DATA_BLOCK "2062_Warning_Data"   // DB2062
{ S7_Optimized_Access := 'FALSE' }
VERSION : 0.1
   VAR
      BTCS_WARNING_WORD_01 : Word;
      BTCS_WARNING_WORD_02 : Word;
      BTCS_WARNING_WORD_03 : Word;
      BTCS_WARNING_WORD_04 : Word;
      BTCS_WARNING_WORD_05 : Word;
      BTCS_WARNING_WORD_06 : Word;
      BTCS_WARNING_WORD_07 : Word;
      BTCS_WARNING_WORD_08 : Word;
      BTCS_WARNING_WORD_09 : Word;
      BTCS_WARNING_WORD_10 : Word;
      BTCS_WARNING_WORD_11 : Word;
      WARNING_PRSNT : Bool;
      "Alarm Tank FPT" : Bool;
      "Alarm Tank P1" : Bool;
      "Alarm Tank S1" : Bool;
      "Alarm Tank P2" : Bool;
      "Alarm Tank S2" : Bool;
      "Alarm Tank P3" : Bool;
      "Alarm Tank S3" : Bool;
      "Alarm Tank P4" : Bool;
      "Alarm Tank S4" : Bool;
      "Alarm Tank P5" : Bool;
      "Alarm Tank S5" : Bool;
      "Alarm Tank P6" : Bool;
      "Alarm Tank S6" : Bool;
      "Alarm Tank APT" : Bool;
      "LS425 FPT Level HIHI" : TON_TIME;
      "LS425 1 Port Level HIHI" : TON_TIME;
      "LS425 1 Starboard Level HIHI" : TON_TIME;
      "PS436 RIO1 Tank Group Pressure HIHI" : TON_TIME;
      "LS425 2 Port Level HIHI" : TON_TIME;
      "LS425 2 Starboard Level HIHI" : TON_TIME;
      "PS436 RIO2 Tank Group Pressure HIHI" : TON_TIME;
      "LS425 3 Port Level HIHI" : TON_TIME;
      "LS425 3 Starboard Level HIHI" : TON_TIME;
      "PS436 RIO3 Tank Group Pressure HIHI" : TON_TIME;
      "LS425 4 Port Level HIHI" : TON_TIME;
      "LS425 4 Starboard Level HIHI" : TON_TIME;
      "PS436 RIO4 Tank Group Pressure HIHI" : TON_TIME;
      "LS425 5 Port Level HIHI" : TON_TIME;
      "LS425 5 Starboard Level HIHI" : TON_TIME;
      "PS436 RIO5 Tank Group Pressure HIHI" : TON_TIME;
      "LS425 6 Port Level HIHI" : TON_TIME;
      "LS425 6 Starboard Level HIHI" : TON_TIME;
      "PS436 RIO6 Tank Group Pressure HIHI" : TON_TIME;
      "LS425 APT Level HIHI" : TON_TIME;
      "PS436 RIO7 Tank Group Pressure HIHI" : TON_TIME;
      "Water Level Override FPT" : Bool;
      "Water Level Override 1P" : Bool;
      "Water Level Override 1S" : Bool;
      "Water Level Override 2P" : Bool;
      "Water Level Override 2S" : Bool;
      "Water Level Override 3P" : Bool;
      "Water Level Override 3S" : Bool;
      "Water Level Override 4P" : Bool;
      "Water Level Override 4S" : Bool;
      "Water Level Override 5P" : Bool;
      "Water Level Override 5S" : Bool;
      "Water Level Override 6P" : Bool;
      "Water Level Override 6S" : Bool;
      "Water Level Override APT" : Bool;
      BTCS_WARNING_WORD_12 : Word;
      BTCS_WARNING_WORD_13 : Word;
      BTCS_WARNING_WORD_14 : Word;
      BTCS_WARNING_WORD_15 : Word;
      BTCS_WARNING_WORD_16 : Word;
      BTCS_WARNING_WORD_17 : Word;
      BTCS_WARNING_WORD_18 : Word;
      "Water Level Override" : Bool;
      "Water Level Override_flag" : Bool;
      "Water Level Override_Aux" : Bool;
   END_VAR
BEGIN
   "LS425 2 Port Level HIHI".PT := T#10s;
   "LS425 2 Starboard Level HIHI".PT := T#10s;
   "PS436 RIO2 Tank Group Pressure HIHI".PT := T#3s;
   "LS425 FPT Level HIHI".PT := T#10s;
   "LS425 1 Port Level HIHI".PT := T#10s;
   "LS425 1 Starboard Level HIHI".PT := T#3s;
END_DATA_BLOCK

DATA_BLOCK "503_WARNING CHCK_DB_2063"   // DB2063
{ S7_Optimized_Access := 'TRUE' }
VERSION : 0.1
// stored: InstanceOfName 503_ALARM CHCK
"503_ALARM CHCK"
BEGIN
END_DATA_BLOCK

DATA_BLOCK "FIT418_2P_ALM_ANALOG_DB"   // DB2064
{ S7_Optimized_Access := 'FALSE' }
VERSION : 0.1
// stored: InstanceOfName 502_ALM_ANALOG
"502_ALM_ANALOG"
BEGIN
END_DATA_BLOCK

DATA_BLOCK "FIT420PORT_ALM_ANALOG_DB"   // DB2065
{ S7_Optimized_Access := 'FALSE' }
VERSION : 0.1
// stored: InstanceOfName 502_ALM_ANALOG
"502_ALM_ANALOG"
BEGIN
END_DATA_BLOCK

DATA_BLOCK "FIT417_2S_ALM_ANALOG_DB"   // DB2066
{ S7_Optimized_Access := 'FALSE' }
VERSION : 0.1
// stored: InstanceOfName 502_ALM_ANALOG
"502_ALM_ANALOG"
BEGIN
END_DATA_BLOCK

DATA_BLOCK "FIT419_ALM_ANALOG_DB"   // DB2067
{ S7_Optimized_Access := 'FALSE' }
VERSION : 0.1
// stored: InstanceOfName 502_ALM_ANALOG
"502_ALM_ANALOG"
BEGIN
END_DATA_BLOCK

DATA_BLOCK "2068_Sys_Status_Data"   // DB2068
{ S7_Optimized_Access := 'TRUE' }
VERSION : 0.1
   VAR
      PORT_GTT_OPEN_FLAG : Bool;   // Confirmed as open after timer
      STBD_GTT_OPEN_FLAG : Bool;   // Confirmed as open after timer
      PORT_GTT_OPEN_TMR : TON_TIME;   // Open timer
      STBD_GTT_OPEN_TMR : TON_TIME;   // Open timer
      SAL_VALID : Bool;   // Validation bit
      SAL_CNF_CHK : Bool;   // Salinity < 1 Confirm bit
      PLS_1 : Bool;   // Pulse bit
      "Not BWT mode Warning" : Bool;
      "LOG BWT" : Bool;   // Tag to log BWT data
      "Times Visibil" : Bool;
      Aux : Struct
         Aux1 : Bool;
         Aux2 : Bool;
         Aux3 : Bool;
      END_STRUCT;
      "Not TANK Activ Warning" : Bool;
      SimulatePuls : Bool;
   END_VAR
BEGIN
   PORT_GTT_OPEN_TMR.PT := T#5s;
   STBD_GTT_OPEN_TMR.PT := T#5s;
END_DATA_BLOCK

DATA_BLOCK "PT415PORT_ALM_ANALOG_DB"   // DB2069
{ S7_Optimized_Access := 'FALSE' }
VERSION : 0.1
// stored: InstanceOfName 502_ALM_ANALOG
"502_ALM_ANALOG"
BEGIN
END_DATA_BLOCK

DATA_BLOCK "PIT424PORT_ALM_ANALOG_DB"   // DB2070
{ S7_Optimized_Access := 'FALSE' }
VERSION : 0.1
// stored: InstanceOfName 502_ALM_ANALOG
"502_ALM_ANALOG"
BEGIN
END_DATA_BLOCK

DATA_BLOCK "TT426PORT_ALM_ANALOG_DB"   // DB2071
{ S7_Optimized_Access := 'FALSE' }
VERSION : 0.1
// stored: InstanceOfName 502_ALM_ANALOG
"502_ALM_ANALOG"
BEGIN
END_DATA_BLOCK

DATA_BLOCK "TT426STR_ALM_ANALOG_DB"   // DB2072
{ S7_Optimized_Access := 'FALSE' }
VERSION : 0.1
// stored: InstanceOfName 502_ALM_ANALOG
"502_ALM_ANALOG"
BEGIN
END_DATA_BLOCK

DATA_BLOCK "TT426PORT_ALM_ANALOG_DB2073"   // DB2073
{ S7_Optimized_Access := 'FALSE' }
VERSION : 0.1
// stored: InstanceOfName 502_ALM_ANALOG
"502_ALM_ANALOG"
BEGIN
END_DATA_BLOCK

DATA_BLOCK "TT426_FPT_ALM_ANALOG_DB"   // DB2074
{ S7_Optimized_Access := 'FALSE' }
VERSION : 0.1
// stored: InstanceOfName 502_ALM_ANALOG
"502_ALM_ANALOG"
BEGIN
END_DATA_BLOCK

DATA_BLOCK "TT426_1P_ALM_ANALOG_DB"   // DB2075
{ S7_Optimized_Access := 'FALSE' }
VERSION : 0.1
// stored: InstanceOfName 502_ALM_ANALOG
"502_ALM_ANALOG"
BEGIN
END_DATA_BLOCK

DATA_BLOCK "TT426_1S_ALM_ANALOG_DB"   // DB2076
{ S7_Optimized_Access := 'FALSE' }
VERSION : 0.1
// stored: InstanceOfName 502_ALM_ANALOG
"502_ALM_ANALOG"
BEGIN
END_DATA_BLOCK

DATA_BLOCK "TT426_3P_ALM_ANALOG_DB"   // DB2077
{ S7_Optimized_Access := 'FALSE' }
VERSION : 0.1
// stored: InstanceOfName 502_ALM_ANALOG
"502_ALM_ANALOG"
BEGIN
END_DATA_BLOCK

DATA_BLOCK "TT426_3S_ALM_ANALOG_DB"   // DB2078
{ S7_Optimized_Access := 'FALSE' }
VERSION : 0.1
// stored: InstanceOfName 502_ALM_ANALOG
"502_ALM_ANALOG"
BEGIN
END_DATA_BLOCK

DATA_BLOCK "TT426_4P_ALM_ANALOG_DB"   // DB2079
{ S7_Optimized_Access := 'FALSE' }
VERSION : 0.1
// stored: InstanceOfName 502_ALM_ANALOG
"502_ALM_ANALOG"
BEGIN
END_DATA_BLOCK

DATA_BLOCK "TT426_4S_ALM_ANALOG_DB"   // DB2080
{ S7_Optimized_Access := 'FALSE' }
VERSION : 0.1
// stored: InstanceOfName 502_ALM_ANALOG
"502_ALM_ANALOG"
BEGIN
END_DATA_BLOCK

DATA_BLOCK "TT426_5P_ALM_ANALOG_DB"   // DB2081
{ S7_Optimized_Access := 'FALSE' }
VERSION : 0.1
// stored: InstanceOfName 502_ALM_ANALOG
"502_ALM_ANALOG"
BEGIN
END_DATA_BLOCK

DATA_BLOCK "TT426_5S_ALM_ANALOG_DB"   // DB2082
{ S7_Optimized_Access := 'FALSE' }
VERSION : 0.1
// stored: InstanceOfName 502_ALM_ANALOG
"502_ALM_ANALOG"
BEGIN
END_DATA_BLOCK

DATA_BLOCK "TT426_6P_ALM_ANALOG_DB"   // DB2083
{ S7_Optimized_Access := 'FALSE' }
VERSION : 0.1
// stored: InstanceOfName 502_ALM_ANALOG
"502_ALM_ANALOG"
BEGIN
END_DATA_BLOCK

DATA_BLOCK "TT426_6S_ALM_ANALOG_DB"   // DB2085
{ S7_Optimized_Access := 'FALSE' }
VERSION : 0.1
// stored: InstanceOfName 502_ALM_ANALOG
"502_ALM_ANALOG"
BEGIN
END_DATA_BLOCK

DATA_BLOCK "TT426_APT_ALM_ANALOG_DB"   // DB2087
{ S7_Optimized_Access := 'FALSE' }
VERSION : 0.1
// stored: InstanceOfName 502_ALM_ANALOG
"502_ALM_ANALOG"
BEGIN
END_DATA_BLOCK

DATA_BLOCK "FIT418_FPT__ALM_ANALOG_DB"   // DB2088
{ S7_Optimized_Access := 'FALSE' }
VERSION : 0.1
// stored: InstanceOfName 502_ALM_ANALOG
"502_ALM_ANALOG"
BEGIN
END_DATA_BLOCK

DATA_BLOCK "FIT418_1P__ALM_ANALOG_DB"   // DB2089
{ S7_Optimized_Access := 'FALSE' }
VERSION : 0.1
// stored: InstanceOfName 502_ALM_ANALOG
"502_ALM_ANALOG"
BEGIN
END_DATA_BLOCK

DATA_BLOCK "FIT417_1S__ALM_ANALOG_DB"   // DB2090
{ S7_Optimized_Access := 'FALSE' }
VERSION : 0.1
// stored: InstanceOfName 502_ALM_ANALOG
"502_ALM_ANALOG"
BEGIN
END_DATA_BLOCK

DATA_BLOCK "FIT418_3P__ALM_ANALOG_DB"   // DB2091
{ S7_Optimized_Access := 'FALSE' }
VERSION : 0.1
// stored: InstanceOfName 502_ALM_ANALOG
"502_ALM_ANALOG"
BEGIN
END_DATA_BLOCK

DATA_BLOCK "FIT417_3S_ALM_ANALOG_DB"   // DB2092
{ S7_Optimized_Access := 'FALSE' }
VERSION : 0.1
// stored: InstanceOfName 502_ALM_ANALOG
"502_ALM_ANALOG"
BEGIN
END_DATA_BLOCK

DATA_BLOCK "FIT418_4P__ALM_ANALOG_DB"   // DB2093
{ S7_Optimized_Access := 'FALSE' }
VERSION : 0.1
// stored: InstanceOfName 502_ALM_ANALOG
"502_ALM_ANALOG"
BEGIN
END_DATA_BLOCK

DATA_BLOCK "FIT417_4S_ALM_ANALOG_DB"   // DB2094
{ S7_Optimized_Access := 'FALSE' }
VERSION : 0.1
// stored: InstanceOfName 502_ALM_ANALOG
"502_ALM_ANALOG"
BEGIN
END_DATA_BLOCK

DATA_BLOCK "FIT418_5P__ALM_ANALOG_DB"   // DB2095
{ S7_Optimized_Access := 'FALSE' }
VERSION : 0.1
// stored: InstanceOfName 502_ALM_ANALOG
"502_ALM_ANALOG"
BEGIN
END_DATA_BLOCK

DATA_BLOCK "FIT417_5S_ALM_ANALOG_DB"   // DB2096
{ S7_Optimized_Access := 'FALSE' }
VERSION : 0.1
// stored: InstanceOfName 502_ALM_ANALOG
"502_ALM_ANALOG"
BEGIN
END_DATA_BLOCK

DATA_BLOCK "FIT418_6P__ALM_ANALOG_DB"   // DB2097
{ S7_Optimized_Access := 'FALSE' }
VERSION : 0.1
// stored: InstanceOfName 502_ALM_ANALOG
"502_ALM_ANALOG"
BEGIN
END_DATA_BLOCK

DATA_BLOCK "FIT417_6S_ALM_ANALOG_DB"   // DB2098
{ S7_Optimized_Access := 'FALSE' }
VERSION : 0.1
// stored: InstanceOfName 502_ALM_ANALOG
"502_ALM_ANALOG"
BEGIN
END_DATA_BLOCK

DATA_BLOCK "FIT417_APT_ALM_ANALOG_DB"   // DB2099
{ S7_Optimized_Access := 'FALSE' }
VERSION : 0.1
// stored: InstanceOfName 502_ALM_ANALOG
"502_ALM_ANALOG"
BEGIN
END_DATA_BLOCK

DATA_BLOCK "O2Analiser_ALM_ANALOG_DB"   // DB2101
{ S7_Optimized_Access := 'FALSE' }
VERSION : 0.1
// stored: InstanceOfName 502_ALM_ANALOG
"502_ALM_ANALOG"
BEGIN
END_DATA_BLOCK

DATA_BLOCK "BWT FPT Ph (426) ALARM"   // DB2103
{ S7_Optimized_Access := 'FALSE' }
VERSION : 0.1
// stored: InstanceOfName 502_ALM_ANALOG
"502_ALM_ANALOG"
BEGIN
END_DATA_BLOCK

DATA_BLOCK "BWT 1P Ph (426) ALARM"   // DB2104
{ S7_Optimized_Access := 'FALSE' }
VERSION : 0.1
// stored: InstanceOfName 502_ALM_ANALOG
"502_ALM_ANALOG"
BEGIN
END_DATA_BLOCK

DATA_BLOCK "BWT 1S Ph (426) ALARM"   // DB2106
{ S7_Optimized_Access := 'FALSE' }
VERSION : 0.1
// stored: InstanceOfName 502_ALM_ANALOG
"502_ALM_ANALOG"
BEGIN
END_DATA_BLOCK

DATA_BLOCK "BWT 2P Ph (426) ALARM"   // DB2107
{ S7_Optimized_Access := 'FALSE' }
VERSION : 0.1
// stored: InstanceOfName 502_ALM_ANALOG
"502_ALM_ANALOG"
BEGIN
END_DATA_BLOCK

DATA_BLOCK "BWT 2S Ph (426) ALARM"   // DB2108
{ S7_Optimized_Access := 'FALSE' }
VERSION : 0.1
// stored: InstanceOfName 502_ALM_ANALOG
"502_ALM_ANALOG"
BEGIN
END_DATA_BLOCK

DATA_BLOCK "BWT 3P Ph (426) ALARM"   // DB2109
{ S7_Optimized_Access := 'FALSE' }
VERSION : 0.1
// stored: InstanceOfName 502_ALM_ANALOG
"502_ALM_ANALOG"
BEGIN
END_DATA_BLOCK

DATA_BLOCK "BWT 3S Ph (426) ALARM"   // DB2111
{ S7_Optimized_Access := 'FALSE' }
VERSION : 0.1
// stored: InstanceOfName 502_ALM_ANALOG
"502_ALM_ANALOG"
BEGIN
END_DATA_BLOCK

DATA_BLOCK "BWT 4P Ph (426) ALARM"   // DB2112
{ S7_Optimized_Access := 'FALSE' }
VERSION : 0.1
// stored: InstanceOfName 502_ALM_ANALOG
"502_ALM_ANALOG"
BEGIN
END_DATA_BLOCK

DATA_BLOCK "BWT 4S Ph (426) ALARM"   // DB2113
{ S7_Optimized_Access := 'FALSE' }
VERSION : 0.1
// stored: InstanceOfName 502_ALM_ANALOG
"502_ALM_ANALOG"
BEGIN
END_DATA_BLOCK

DATA_BLOCK "BWT 5P Ph (426) ALARM"   // DB2114
{ S7_Optimized_Access := 'FALSE' }
VERSION : 0.1
// stored: InstanceOfName 502_ALM_ANALOG
"502_ALM_ANALOG"
BEGIN
END_DATA_BLOCK

DATA_BLOCK "BWT 5S Ph (426) ALARM"   // DB2116
{ S7_Optimized_Access := 'FALSE' }
VERSION : 0.1
// stored: InstanceOfName 502_ALM_ANALOG
"502_ALM_ANALOG"
BEGIN
END_DATA_BLOCK

DATA_BLOCK "BWT 6P Ph (426) ALARM"   // DB2117
{ S7_Optimized_Access := 'FALSE' }
VERSION : 0.1
// stored: InstanceOfName 502_ALM_ANALOG
"502_ALM_ANALOG"
BEGIN
END_DATA_BLOCK

DATA_BLOCK "BWT 6S Ph (426) ALARM"   // DB2118
{ S7_Optimized_Access := 'FALSE' }
VERSION : 0.1
// stored: InstanceOfName 502_ALM_ANALOG
"502_ALM_ANALOG"
BEGIN
END_DATA_BLOCK

DATA_BLOCK "BWT APT Ph (426) ALARM"   // DB2119
{ S7_Optimized_Access := 'FALSE' }
VERSION : 0.1
// stored: InstanceOfName 502_ALM_ANALOG
"502_ALM_ANALOG"
BEGIN
END_DATA_BLOCK

DATA_BLOCK "BWT FPT DO (426) ALARM"   // DB2120
{ S7_Optimized_Access := 'FALSE' }
VERSION : 0.1
// stored: InstanceOfName 502_ALM_ANALOG
"502_ALM_ANALOG"
BEGIN
END_DATA_BLOCK

DATA_BLOCK "BWT 1P DO (426) ALARM"   // DB2121
{ S7_Optimized_Access := 'FALSE' }
VERSION : 0.1
// stored: InstanceOfName 502_ALM_ANALOG
"502_ALM_ANALOG"
BEGIN
END_DATA_BLOCK

DATA_BLOCK "BWT 1S DO (426) ALARM"   // DB2122
{ S7_Optimized_Access := 'FALSE' }
VERSION : 0.1
// stored: InstanceOfName 502_ALM_ANALOG
"502_ALM_ANALOG"
BEGIN
END_DATA_BLOCK

DATA_BLOCK "BWT 2P DO (426) ALARM"   // DB2123
{ S7_Optimized_Access := 'FALSE' }
VERSION : 0.1
// stored: InstanceOfName 502_ALM_ANALOG
"502_ALM_ANALOG"
BEGIN
END_DATA_BLOCK

DATA_BLOCK "BWT 2S DO (426) ALARM"   // DB2124
{ S7_Optimized_Access := 'FALSE' }
VERSION : 0.1
// stored: InstanceOfName 502_ALM_ANALOG
"502_ALM_ANALOG"
BEGIN
END_DATA_BLOCK

DATA_BLOCK "BWT 3P DO (426) ALARM"   // DB2125
{ S7_Optimized_Access := 'FALSE' }
VERSION : 0.1
// stored: InstanceOfName 502_ALM_ANALOG
"502_ALM_ANALOG"
BEGIN
END_DATA_BLOCK

DATA_BLOCK "BWT 3S DO (426) ALARM"   // DB2126
{ S7_Optimized_Access := 'FALSE' }
VERSION : 0.1
// stored: InstanceOfName 502_ALM_ANALOG
"502_ALM_ANALOG"
BEGIN
END_DATA_BLOCK

DATA_BLOCK "BWT 4P DO (426) ALARM"   // DB2127
{ S7_Optimized_Access := 'FALSE' }
VERSION : 0.1
// stored: InstanceOfName 502_ALM_ANALOG
"502_ALM_ANALOG"
BEGIN
END_DATA_BLOCK

DATA_BLOCK "BWT 4S DO (426) ALARM"   // DB2128
{ S7_Optimized_Access := 'FALSE' }
VERSION : 0.1
// stored: InstanceOfName 502_ALM_ANALOG
"502_ALM_ANALOG"
BEGIN
END_DATA_BLOCK

DATA_BLOCK "BWT 5P DO (426) ALARM"   // DB2129
{ S7_Optimized_Access := 'FALSE' }
VERSION : 0.1
// stored: InstanceOfName 502_ALM_ANALOG
"502_ALM_ANALOG"
BEGIN
END_DATA_BLOCK

DATA_BLOCK "BWT 5S DO (426) ALARM"   // DB2130
{ S7_Optimized_Access := 'FALSE' }
VERSION : 0.1
// stored: InstanceOfName 502_ALM_ANALOG
"502_ALM_ANALOG"
BEGIN
END_DATA_BLOCK

DATA_BLOCK "BWT 6P DO (426) ALARM"   // DB2131
{ S7_Optimized_Access := 'FALSE' }
VERSION : 0.1
// stored: InstanceOfName 502_ALM_ANALOG
"502_ALM_ANALOG"
BEGIN
END_DATA_BLOCK

DATA_BLOCK "BWT 6S DO (426) ALARM"   // DB2132
{ S7_Optimized_Access := 'FALSE' }
VERSION : 0.1
// stored: InstanceOfName 502_ALM_ANALOG
"502_ALM_ANALOG"
BEGIN
END_DATA_BLOCK

DATA_BLOCK "BWT APT DO (426) ALARM"   // DB2133
{ S7_Optimized_Access := 'FALSE' }
VERSION : 0.1
// stored: InstanceOfName 502_ALM_ANALOG
"502_ALM_ANALOG"
BEGIN
END_DATA_BLOCK

DATA_BLOCK "FIT420_FPT_ALM_ANALOG_DB"   // DB2201
{ S7_Optimized_Access := 'FALSE' }
VERSION : 0.1
// stored: InstanceOfName 502_ALM_ANALOG
"502_ALM_ANALOG"
BEGIN
END_DATA_BLOCK

DATA_BLOCK "FIT420_1P_ALM_ANALOG_DB"   // DB2202
{ S7_Optimized_Access := 'FALSE' }
VERSION : 0.1
// stored: InstanceOfName 502_ALM_ANALOG
"502_ALM_ANALOG"
BEGIN
END_DATA_BLOCK

DATA_BLOCK "FIT420_1S_ALM_ANALOG_DB"   // DB2203
{ S7_Optimized_Access := 'FALSE' }
VERSION : 0.1
// stored: InstanceOfName 502_ALM_ANALOG
"502_ALM_ANALOG"
BEGIN
END_DATA_BLOCK

DATA_BLOCK "FIT420_3P_ALM_ANALOG_DB"   // DB2204
{ S7_Optimized_Access := 'FALSE' }
VERSION : 0.1
// stored: InstanceOfName 502_ALM_ANALOG
"502_ALM_ANALOG"
BEGIN
END_DATA_BLOCK

DATA_BLOCK "FIT420_3S_ALM_ANALOG_DB"   // DB2205
{ S7_Optimized_Access := 'FALSE' }
VERSION : 0.1
// stored: InstanceOfName 502_ALM_ANALOG
"502_ALM_ANALOG"
BEGIN
END_DATA_BLOCK

DATA_BLOCK "FIT420_4P_ALM_ANALOG_DB"   // DB2206
{ S7_Optimized_Access := 'FALSE' }
VERSION : 0.1
// stored: InstanceOfName 502_ALM_ANALOG
"502_ALM_ANALOG"
BEGIN
END_DATA_BLOCK

DATA_BLOCK "FIT420_4S_ALM_ANALOG_DB"   // DB2207
{ S7_Optimized_Access := 'FALSE' }
VERSION : 0.1
// stored: InstanceOfName 502_ALM_ANALOG
"502_ALM_ANALOG"
BEGIN
END_DATA_BLOCK

DATA_BLOCK "FIT420_5P_ALM_ANALOG_DB"   // DB2208
{ S7_Optimized_Access := 'FALSE' }
VERSION : 0.1
// stored: InstanceOfName 502_ALM_ANALOG
"502_ALM_ANALOG"
BEGIN
END_DATA_BLOCK

DATA_BLOCK "FIT420_5S_ALM_ANALOG_DB"   // DB2209
{ S7_Optimized_Access := 'FALSE' }
VERSION : 0.1
// stored: InstanceOfName 502_ALM_ANALOG
"502_ALM_ANALOG"
BEGIN
END_DATA_BLOCK

DATA_BLOCK "FIT420_6P_ALM_ANALOG_DB"   // DB2210
{ S7_Optimized_Access := 'FALSE' }
VERSION : 0.1
// stored: InstanceOfName 502_ALM_ANALOG
"502_ALM_ANALOG"
BEGIN
END_DATA_BLOCK

DATA_BLOCK "FIT420_6S_ALM_ANALOG_DB"   // DB2211
{ S7_Optimized_Access := 'FALSE' }
VERSION : 0.1
// stored: InstanceOfName 502_ALM_ANALOG
"502_ALM_ANALOG"
BEGIN
END_DATA_BLOCK

DATA_BLOCK "FIT420_APT_ALM_ANALOG_DB"   // DB2212
{ S7_Optimized_Access := 'FALSE' }
VERSION : 0.1
// stored: InstanceOfName 502_ALM_ANALOG
"502_ALM_ANALOG"
BEGIN
END_DATA_BLOCK

DATA_BLOCK "PT415_FPT_ALM_ANALOG_DB"   // DB2213
{ S7_Optimized_Access := 'FALSE' }
VERSION : 0.1
// stored: InstanceOfName 502_ALM_ANALOG
"502_ALM_ANALOG"
BEGIN
END_DATA_BLOCK

DATA_BLOCK "PT415_1P_ALM_ANALOG_DB"   // DB2214
{ S7_Optimized_Access := 'FALSE' }
VERSION : 0.1
// stored: InstanceOfName 502_ALM_ANALOG
"502_ALM_ANALOG"
BEGIN
END_DATA_BLOCK

DATA_BLOCK "PT415_RIO3_ALM_ANALOG_DB"   // DB2215
{ S7_Optimized_Access := 'FALSE' }
VERSION : 0.1
// stored: InstanceOfName 502_ALM_ANALOG
"502_ALM_ANALOG"
BEGIN
END_DATA_BLOCK

DATA_BLOCK "PT415_RIO4_ALM_ANALOG_DB"   // DB2216
{ S7_Optimized_Access := 'FALSE' }
VERSION : 0.1
// stored: InstanceOfName 502_ALM_ANALOG
"502_ALM_ANALOG"
BEGIN
END_DATA_BLOCK

DATA_BLOCK "PT415_RIO5_ALM_ANALOG_DB"   // DB2217
{ S7_Optimized_Access := 'FALSE' }
VERSION : 0.1
// stored: InstanceOfName 502_ALM_ANALOG
"502_ALM_ANALOG"
BEGIN
END_DATA_BLOCK

DATA_BLOCK "PT415_RIO6_ALM_ANALOG_DB"   // DB2218
{ S7_Optimized_Access := 'FALSE' }
VERSION : 0.1
// stored: InstanceOfName 502_ALM_ANALOG
"502_ALM_ANALOG"
BEGIN
END_DATA_BLOCK

DATA_BLOCK "PIT424_RIO1_ALM_ANALOG_DB"   // DB2219
{ S7_Optimized_Access := 'FALSE' }
VERSION : 0.1
// stored: InstanceOfName 502_ALM_ANALOG
"502_ALM_ANALOG"
BEGIN
END_DATA_BLOCK

DATA_BLOCK "PIT424_RIO3_ALM_ANALOG_DB"   // DB2220
{ S7_Optimized_Access := 'FALSE' }
VERSION : 0.1
// stored: InstanceOfName 502_ALM_ANALOG
"502_ALM_ANALOG"
BEGIN
END_DATA_BLOCK

DATA_BLOCK "PIT424_RIO4_ALM_ANALOG_DB"   // DB2221
{ S7_Optimized_Access := 'FALSE' }
VERSION : 0.1
// stored: InstanceOfName 502_ALM_ANALOG
"502_ALM_ANALOG"
BEGIN
END_DATA_BLOCK

DATA_BLOCK "PIT424_RIO5_ALM_ANALOG_DB"   // DB2222
{ S7_Optimized_Access := 'FALSE' }
VERSION : 0.1
// stored: InstanceOfName 502_ALM_ANALOG
"502_ALM_ANALOG"
BEGIN
END_DATA_BLOCK

DATA_BLOCK "PIT424_RIO6_ALM_ANALOG_DB"   // DB2223
{ S7_Optimized_Access := 'FALSE' }
VERSION : 0.1
// stored: InstanceOfName 502_ALM_ANALOG
"502_ALM_ANALOG"
BEGIN
END_DATA_BLOCK

DATA_BLOCK "PIT424_RIO7_ALM_ANALOG_DB"   // DB2224
{ S7_Optimized_Access := 'FALSE' }
VERSION : 0.1
// stored: InstanceOfName 502_ALM_ANALOG
"502_ALM_ANALOG"
BEGIN
END_DATA_BLOCK

DATA_BLOCK "PT415_RIO7_ALM_ANALOG_DB"   // DB2225
{ S7_Optimized_Access := 'FALSE' }
VERSION : 0.1
// stored: InstanceOfName 502_ALM_ANALOG
"502_ALM_ANALOG"
BEGIN
END_DATA_BLOCK

DATA_BLOCK "LT422 FPT  TANK LEVEL ALARM"   // DB2226
{ S7_Optimized_Access := 'FALSE' }
VERSION : 0.1
// stored: InstanceOfName 502_ALM_ANALOG
"502_ALM_ANALOG"
BEGIN
END_DATA_BLOCK

DATA_BLOCK "LT422 1P  TANK LEVEL ALARM"   // DB2227
{ S7_Optimized_Access := 'FALSE' }
VERSION : 0.1
// stored: InstanceOfName 502_ALM_ANALOG
"502_ALM_ANALOG"
BEGIN
END_DATA_BLOCK

DATA_BLOCK "LT421 1S  TANK LEVEL ALARM"   // DB2228
{ S7_Optimized_Access := 'FALSE' }
VERSION : 0.1
// stored: InstanceOfName 502_ALM_ANALOG
"502_ALM_ANALOG"
BEGIN
END_DATA_BLOCK

DATA_BLOCK "LT422 2P  TANK LEVEL ALARM"   // DB2229
{ S7_Optimized_Access := 'FALSE' }
VERSION : 0.1
// stored: InstanceOfName 502_ALM_ANALOG
"502_ALM_ANALOG"
BEGIN
END_DATA_BLOCK

DATA_BLOCK "LT421 2S  TANK LEVEL ALARM"   // DB2230
{ S7_Optimized_Access := 'FALSE' }
VERSION : 0.1
// stored: InstanceOfName 502_ALM_ANALOG
"502_ALM_ANALOG"
BEGIN
END_DATA_BLOCK

DATA_BLOCK "LT422 3P  TANK LEVEL ALARM"   // DB2231
{ S7_Optimized_Access := 'FALSE' }
VERSION : 0.1
// stored: InstanceOfName 502_ALM_ANALOG
"502_ALM_ANALOG"
BEGIN
END_DATA_BLOCK

DATA_BLOCK "LT421 3S  TANK LEVEL ALARM"   // DB2232
{ S7_Optimized_Access := 'FALSE' }
VERSION : 0.1
// stored: InstanceOfName 502_ALM_ANALOG
"502_ALM_ANALOG"
BEGIN
END_DATA_BLOCK

DATA_BLOCK "LT422 4P  TANK LEVEL ALARM"   // DB2233
{ S7_Optimized_Access := 'FALSE' }
VERSION : 0.1
// stored: InstanceOfName 502_ALM_ANALOG
"502_ALM_ANALOG"
BEGIN
END_DATA_BLOCK

DATA_BLOCK "LT421 4S  TANK LEVEL ALARM"   // DB2234
{ S7_Optimized_Access := 'FALSE' }
VERSION : 0.1
// stored: InstanceOfName 502_ALM_ANALOG
"502_ALM_ANALOG"
BEGIN
END_DATA_BLOCK

DATA_BLOCK "LT422 5P  TANK LEVEL ALARM"   // DB2235
{ S7_Optimized_Access := 'FALSE' }
VERSION : 0.1
// stored: InstanceOfName 502_ALM_ANALOG
"502_ALM_ANALOG"
BEGIN
END_DATA_BLOCK

DATA_BLOCK "LT421 5S  TANK LEVEL ALARM"   // DB2236
{ S7_Optimized_Access := 'FALSE' }
VERSION : 0.1
// stored: InstanceOfName 502_ALM_ANALOG
"502_ALM_ANALOG"
BEGIN
END_DATA_BLOCK

DATA_BLOCK "LT422 6P  TANK LEVEL ALARM"   // DB2237
{ S7_Optimized_Access := 'FALSE' }
VERSION : 0.1
// stored: InstanceOfName 502_ALM_ANALOG
"502_ALM_ANALOG"
BEGIN
END_DATA_BLOCK

DATA_BLOCK "LT421 6S  TANK LEVEL ALARM"   // DB2238
{ S7_Optimized_Access := 'FALSE' }
VERSION : 0.1
// stored: InstanceOfName 502_ALM_ANALOG
"502_ALM_ANALOG"
BEGIN
END_DATA_BLOCK

DATA_BLOCK "LT422 APT  TANK LEVEL ALARM"   // DB2239
{ S7_Optimized_Access := 'FALSE' }
VERSION : 0.1
// stored: InstanceOfName 502_ALM_ANALOG
"502_ALM_ANALOG"
BEGIN
END_DATA_BLOCK

DATA_BLOCK "BTCS_ALARM_CHK_DB"   // DB2500
{ S7_Optimized_Access := 'TRUE' }
VERSION : 0.1
// stored: InstanceOfName 503_ALARM CHCK
"503_ALARM CHCK"
BEGIN
END_DATA_BLOCK

// folder: 2000 - 2999 BTCS System/2080 - 2089 HMI Handling

DATA_BLOCK "2084_Setpoints"   // DB2084
TITLE = Setpoints Data
{ S7_Optimized_Access := 'TRUE' }
AUTHOR : JRS
VERSION : 0.1
// Setpoints data area
   VAR RETAIN
      PIT415_LoLo : Real := 0.4;
      PIT415_Lo : Real := 0.5;
      PIT415_Hi : Real := 5.5;
      PIT415_HiHi : Real := 6.0;
      PIT424_LoLo : Real := 0.0;
      PIT424_Lo : Real := 0.0;
      PIT424_Hi : Real := 80.0;
      PIT424_HiHi : Real := 85.0;
      FIT417_LoLo : Real := -85.0;
      FIT417_Lo : Real := -75.0;
      FIT417_Hi : Real := 400.0;
      FIT417_HiHi : Real := 450.0;
      FIT418_LoLo : Real := 0.0;
      FIT418_Lo : Real := 0.0;
      FIT418_Hi : Real := 400.0;
      FIT418_HiHi : Real := 450.0;
      FIT419_LoLo : Real := 0.0;
      FIT419_Lo : Real := 0.0;
      FIT419_Hi : Real := 350.0;
      FIT419_HiHi : Real := 400.0;
      FIT420_LoLo : Real := 0.0;
      FIT420_Lo : Real := 0.0;
      FIT420_Hi : Real := 350.0;
      FIT420_HiHi : Real := 400.0;
      LT422_Lo : Real := 50.0;
      LT422_Hi : Real := 98.0;
      LT421_Lo : Real := 50.0;
      LT421_Hi : Real := 98.0;
      TT436_Hi : Real := 75.0;
      TT436_HiHi : Real := 85.0;
      DO_SP : Real := 22.0;
      PH_SP : Real := 6.5;
      "TX426 Port PH Lo" : Real := 1.0;
      "TX426 Port PH High" : Real := 20.0;
      "TX428 Port DO Lo" : Real := 0.0;
      "TX428 Port DO High" : Real := 20.0;
      "TX425 Star PH Lo" : Real := 1.0;
      "TX425 Star PH High" : Real := 50.0;
      "TX427 Star DO Lo" : Real := 0.0;
      "TX427 Star DO High" : Real := 20.0;
   END_VAR
   VAR
      "Conf O2 Level Lo" : Real := 10.0;
      "Conf O2 Level Lo Lo" : Real := 16.0;
   END_VAR
BEGIN
END_DATA_BLOCK

DATA_BLOCK "2086_Times"   // DB2086
TITLE = Times Data
{ S7_Optimized_Access := 'TRUE' }
AUTHOR : JRS
VERSION : 0.1
// Times data area
   VAR RETAIN
      DEOX_PRE_GTT_OPN_DLY : Time := T#15S;   // Sequence step delay time
      DEOX_PRE_GTT_CLS_DLY : Time := T#15S;   // Sequence step delay time
      REOX_PRE_GTT_OPN_DLY : Time := T#15S;   // Sequence step delay time
      REOX_PRE_GTT_CLS_DLY : Time := T#15S;   // Sequence step delay time
      AT_DEOX_CNF_TIME : Time := T#1M;   // Sequence step delay time
      AT_REOX_CNF_TIME : Time := T#1M;   // Sequence step delay time
      CV422_FPT_MAX_TRVL_TIME : Time := T#3M;
      CV422_1P_MAX_TRVL_TIME : Time := T#3M;
      CV421_1S_MAX_TRVL_TIME : Time := T#3M;
      CV422_2P_MAX_TRVL_TIME : Time := T#3M;   // Maximum valve travel time
      CV421_2S_MAX_TRVL_TIME : Time := T#3M;   // Maximum valve travel time
      CV422_3P_MAX_TRVL_TIME : Time := T#3M;
      CV421_3S_MAX_TRVL_TIME : Time := T#3M;
      CV422_4P_MAX_TRVL_TIME : Time := T#3M;
      CV421_4S_MAX_TRVL_TIME : Time := T#3M;
      CV422_5P_MAX_TRVL_TIME : Time := T#3M;
      CV421_5S_MAX_TRVL_TIME : Time := T#3M;
      CV422_6P_MAX_TRVL_TIME : Time := T#3M;
      CV421_6S_MAX_TRVL_TIME : Time := T#3M;
      CV422_APT_MAX_TRVL_TIME : Time := T#3M;
      "TT426_PORT_Alarm Delay" : Time := T#5S;
      "TT426_STAR_Alarm Delay" : Time := T#5S;
      "FIT418PORT Alarm Delay" : Time := T#10S;
      "FIT420PORT Alarm Delay" : Time := T#10S;
      "FIT417STAR Alarm Delay" : Time := T#10S;
      "FIT419STAR Alarm Delay" : Time := T#10S;
      "PT415 Alarm Delay" : Time := T#30S;
      "PIT424 Alarm Delay" : Time := T#30S;
      "LS425 Port Alarm Delay" : Time := T#30S;
      "LS425 Star Alarm Delay" : Time := T#30S;
      "PS436 Alarm Delay" : Time := T#30S;
      "TIMER RST Supres" : Bool := FALSE;   // TIMER RST Supres
      "Tank Alarm Reset Time" : Time := T#1M;
      "Alarm Enable Delay" : Time := T#1S;
      "LT422 Alarm Delay" : Time := T#30S;
   END_VAR
   VAR
      "LT421 Alarm Delay" : Time := T#30S;
      "Stage Warning" : Time := T#3MS;   // Warning to start IGG befor De-Ox and GCU before Re-Ox
   END_VAR
BEGIN
END_DATA_BLOCK

// folder: 2000 - 2999 BTCS System/2100 - 2199 Automatic Sequencing

DATA_BLOCK "2100_AUTO_SEQ_DB"   // DB2100
TITLE = Automatic Sequence Data Area
{ S7_Optimized_Access := 'TRUE' }
AUTHOR : JRS
VERSION : 0.1
// Primary data area for the automatic sequence related data
   VAR
      INI_DN : Bool := false;   // 1 = Block has started & set defaults, 0 = Not
      SEQ_RNG : Bool := false;   // 1 = Sequence running, 0 = Not
   END_VAR
BEGIN
END_DATA_BLOCK

DATA_BLOCK "2102_TIME_CALCS_DB"   // DB2102
TITLE = TTime Calculations Data Area
{ S7_Optimized_Access := 'TRUE' }
AUTHOR : JRS
VERSION : 0.1
// Primary data area for time calculations
   VAR
      Voyage_TIME_days : Int;
      Voyage_TIME_hours : Int;
      Voyage_TIME_min : Int;
      Voyage_TIME_shorter_min : Int;   // Voyage time shorter than BWT sequence
      Voyage_TIME_shorter_hours : Int;
      Voyage_TIME_invalid : Bool;   // Voyage time shorter than BWT sequence
      Voyage_TIME_remaining_h : Int;
      Voyage_TIME_remaining_m : Int;
      "PRE-DWEL_Warning 1" : Bool;
      "PRE-DWEL_Warning 2" : Bool;
      "PRE-DWEL_Warning 3" : Bool;
      "PRE-DWEL_Warning Min 1" : Int := 1;
      "PRE-DWEL_Warning Min 2" : Int := 2;
      "PRE-DWEL_Warning Min 3" : Int := 3;
      "PRE-DWEL_Warning Reset 1" : Bool;
      "PRE-DWEL_Warning Reset 2" : Bool;
      "PRE-DWEL_Warning Reset 3" : Bool;
      "PRE-DWEL_Warning Reset Aux 1" : Bool;
      "PRE-DWEL_Warning Reset Aux 2" : Bool;
      "PRE-DWEL_Warning Reset Aux 3" : Bool;
      "PRE-DWEL_Warning Puls Aux 1" : Bool;
      "PRE-DWEL_Warning Puls Aux 2" : Bool;
      "PRE-DWEL_Warning Puls Aux 3" : Bool;
      "PRE-DWEL_Warning Puls 1" : Bool;
      "PRE-DWEL_Warning Puls 2" : Bool;
      "PRE-DWEL_Warning Puls 3" : Bool;
      PRE_DWELL_MINS : Int := 0;   // Total time in minutes
      PRE_DWELL_HRS : Int;
      DE_OX_MINS : Int;   // Total time in minutes
      DE_OX_SP_MINS : Int;   // Total time in minutes
      DWELL_MINS : Int;   // Total time in minutes
      RE_OX_MINS : Int;   // Total time in minutes
      RE_OX_SP_MINS : Int;   // Total time in minutes
      POST_DWELL_MINS : Int;   // Total time in minutes
      TOT_SEQ_MINS : Int;   // Total time in minutes
      TOT_SEQ_DAYS : Real;
      "PRE-DWEL HOURS REMNG" : Int;   // Time remaining until the start of DeOx is required
      "PRE-DWEL MINS REMNG" : Int;
      SCNDS_COUNT : Int;   // Seconds Count
      MNTS_COUNT : Int;
      TIMES_VALID : Bool := false;   // 1 = Input times valid, 0 = Not
      INTO_RNG_PLS : Bool := false;   // Pulse bit
      CLK_PLS : Bool := false;   // Pulse bit
      PRE_DWELL_TMR_DN : Bool := false;   // Count down done
      DE_OX_TMR_DN : Bool := false;   // Count down done
      DE_OX_SP_TMR_DN : Bool;   // Count down done
      DWELL_TMR_DN : Bool := false;   // Count down done
      RE_OX_TMR_DN : Bool := false;   // Count down done
      RE_OX_SP_TMR_DN : Bool;   // Count down done
      POST_DWELL_TMR_DN : Bool := false;   // Count down done
      PRE_DWELL_MINS_RMNG : Int := 0;   // Total time remaining in minutes
      DE_OX_MINS_RMNG : Int;   // Total time remaining in minutes
      DE_OX_SP_MINS_RMNG : Int;   // Total time remaining in minutes
      DWELL_MINS_RMNG : Int;   // Total time remaining in minutes
      RE_OX_MINS_RMNG : Int;   // Total time remaining in minutes
      RE_OX_SP_MINS_RMNG : Int;   // Total time remaining in minutes
      POST_DWELL_MINS_RMNG : Int;   // Total time remaining in minutes
      TOT_SEQ_MINS_RMNG : Int;   // Total time remaining in minutes
      TOT_SEQ_HRS_RMNG : Int;   // Total time remaining in hours
      Voyage_TIME : CTD_INT;
      PRE_DWELL_CNTR : CTD_INT;   // Counter
   END_VAR
   VAR RETAIN
      DE_OX_CNTR : CTD_INT;   // Counter
      DE_OX_SP_CNTR : CTD_INT;   // Counter
      DWELL_CNTR : CTD_INT;   // Counter
      RE_OX_CNTR : CTD_INT;   // Counter
      RE_OX_SP_CNTR : CTD_INT;   // Counter
      POST_DWELL_CNTR : CTD_INT;   // Counter
      MINUTE : Bool;   // Full minute reached
   END_VAR
   VAR
      HOUR : Bool;   // Full hour reached
      MIN_PLS : Bool;   // Pulse bit
      Hour_PLS : Bool;
      "60X boost" : Bool;   // Times accelerated 60 times
      ONE_SEC_PULS : Bool;
      Voyage_Popup_ACC : Int;   // Accumulated Seconds for Voyage Popup
      Time_To_Treatment : Int;   // Time Until Treatment Required
      PHASE_DIFFERECE_MNS : Int;
      "PHASE_DIFFERECE_MNS_REMNG_De-Ox" : Int;
      "DE_OX_MINS_RMNG_Scnd GROUP" : Int;
      "PHASE_DIFFERECE_MNS_REMNG_Re-Ox" : Int;
      "DE_OX_SP_MINS_RMNG_Scnd GROUP" : Int;
      "DWELL_MINS_RMNG_Scnd GROUP" : Int;
      "RE_OX_MINS_RMNG_Scnd GROUP" : Int;
      "RE_OX_SP_MINS_RMNG_Scnd GROUP" : Int;
   END_VAR
BEGIN
END_DATA_BLOCK

DATA_BLOCK "Sequence Times_DB"   // DB2105
{ S7_Optimized_Access := 'TRUE' }
VERSION : 0.1
// stored: InstanceOfName Sequence Times
"Sequence Times"
BEGIN
END_DATA_BLOCK

DATA_BLOCK "2110_BTCS_CNTRL_DB"   // DB2110
TITLE = Barge Tank Control System Data Area
{ S7_Optimized_Access := 'TRUE' }
AUTHOR : JRS
VERSION : 0.1
// Primary data area for barge tank control related data
   VAR
      BTCS_STATE : Int := 0;   // 0=Init, 1=PreDwell, 2=DeOx, 3=Dwell, 4=ReOx, 5 = PostDwell & Done, 6=SD
      BTCS_STEP : Int := 0;   // BTCS Sequence step number
      PORT_TANK_STS : Bool := 1;   // 0 = Isolated, 1 = Active, add as needed
      STBD_TANK_STS : Bool := 1;   // 0 = Isolated, 1 = Active, add as needed
      VNT_VLV_CNTRL_PRSNT : Bool;   // 1 = Vent Valve Control Fitted, 0 = Not
      PRE_DWELL_HRS : Int := 18;   // Pre-dwell time
      DE_OX_HRS : Int := 10;   // De-oxygenate time
      DE_OX_SP_HRS : Int := 2;   // Minimum run at setpoint + DeOx
      DWELL_HRS : Int := 60;   // Dwell time
      RE_OX_HRS : Int := 6;   // Re-oxygenate time
      RE_OX_SP_HRS : Int := 2;   // Minimum run at setpoint + ReOx
      POST_DWELL_HRS : Int := 12;   // Post-dwell time
      PRE_DWELL_MINS : Int := 0;   // Pre-dwell time
      DE_OX_MINS : Int := 0;   // De-oxygenate time
      DE_OX_SP_MINS : Int := 0;   // Minimum run at setpoint + DeOx
      DWELL_MINS : Int := 0;   // Dwell time
      RE_OX_MINS : Int := 0;   // Re-oxygenate time
      RE_OX_SP_MINS : Int := 0;   // Minimum run at setpoint + ReOx
      POST_DWELL_MINS : Int := 0;   // Post-dwell time
      TOT_SEQ_HRS : Int := 0;   // Total sequence hours
      TOT_SEQ_MINS : Int := 0;   // Total sequence minutes
      RMNG_SEQ_HRS : Int := 0;   // Remaining sequence hours
      RMNG_SEQ_MINS : Int := 0;   // Remaining sequence minutes
      MSTR_RST_PLS : TP_TIME;   // Master Reset Pulse
      START_SEQ : Bool;   // Accept timings and run
      STOP_SEQ : Bool;   // Stop and shutdown sequence
      STOP_MSTR_FLG : Bool;   // Master stop sequence flag
      STOP_PLS : Bool;   // Pulse bit
      RESET_ALL : Bool;   // Master reset from HMI
      INTO_BTCS_PLS : Bool;   // Pulse bit
      OUT_BTCS_PLS : Bool;   // Pulse bit
      RE_OX_DN : Bool;   // Re-oxygenate done
      VNT_VLV_STS_OK : Bool;   // Vent valves as expected for active tanks
      GTT_VLV_STS_OK : Bool;   // GTT valves as expected for active tanks
      O2_AT_DEOX : Bool;   // Active tanks O2 level at de-ox
      O2_AT_REOX : Bool;   // Active tanks O2 level at re-ox
      O2_AT_DEOX_CNFMD : Bool;   // Active tanks O2 level at de-ox confirmed
      O2_AT_REOX_CNFMD : Bool;   // Active tanks O2 level at re-ox confirmed
      TIME_DLY_STEP_45 : TON_TIME;   // Sequence delay timer
      TIME_DLY_STEP_80 : TON_TIME;   // Sequence delay timer
      TIME_DLY_STEP_145 : TON_TIME;   // Sequence delay timer
      TIME_DLY_STEP_180 : TON_TIME;   // Sequence delay timer
      O2_AT_DEOX_TMR : TON_TIME;   // Confirmation of O2 at de-ox level
      O2_AT_REOX_TMR : TON_TIME;   // Confirmation of O2 at re-ox level
      PHASE_DIFFERECE_HRS : Int;
      PHASE_DIFFERECE_MNS : Int;
      "O2_AT_DEOX_CNFMD_Scnd GROUP" : Bool;
      Auxiliary : Struct
         "Aux 1" : Bool;
      END_STRUCT;
   END_VAR
BEGIN
   MSTR_RST_PLS.PT := T#100ms;
   TIME_DLY_STEP_45.PT := T#15s;
   O2_AT_DEOX_TMR.PT := T#60s;
   TIME_DLY_STEP_80.PT := T#30s;
   TIME_DLY_STEP_145.PT := T#15s;
   O2_AT_REOX_TMR.PT := T#60s;
   TIME_DLY_STEP_180.PT := T#30s;
END_DATA_BLOCK

DATA_BLOCK "2115_VOYAGE_TIME_DAYS"   // DB2115
{ S7_Optimized_Access := 'TRUE' }
VERSION : 0.1
   VAR
      VOYAGE_DAYS : Real;
      VOYAGE_HOURS : Real;
      VOYAGE_MINUTE : Real;
   END_VAR
BEGIN
END_DATA_BLOCK

// folder: 300 - 499 Counter and Timer DBs

DATA_BLOCK "300_AUT_SEQ_TMRS_DB"   // DB300
TITLE = Auto Sequence Timers Data
{ S7_Optimized_Access := 'TRUE' }
AUTHOR : JRS